(* Logix 5000 project; controller NWGG 1756-L72 rev 35.12; software revision 35.00; part 8 of 19 *)
(* tags used below, declared in another part *)
   _700_AIR_GA : ALIAS FOR I8.3;
   _700_METER : ALIAS FOR I8.2;
   _700_TREAT : ALIAS FOR I7.3;
   _700G_13_CL : ALIAS FOR B21[70].1;
   _700G_13_OP : ALIAS FOR B21[70].0;
   _700G_CLOSE : ALIAS FOR O12.9;
   _700G_OPEN : ALIAS FOR O12.8;
   _701_AIR_GA : ALIAS FOR I8.5;
   _701_FB : ALIAS FOR B21[1].3;
   _701_K_TREA : ALIAS FOR I8.0;
   _701_METER : ALIAS FOR I8.4;
   _701_RB : ALIAS FOR B21[1].4;
   _701_REV_CN : ALIAS FOR C5[3];
   _701_STP : ALIAS FOR B21[1].2;
   _701F_HPB : ALIAS FOR B21[1].0;
   _701F_M : ALIAS FOR O25[10].11;
   _701F_OFF_T : ALIAS FOR T22[1];
   _701G_CLOSE : ALIAS FOR B21[71].13;
   _701G_OPEN : ALIAS FOR B21[71].12;
   _701MR : ALIAS FOR O25[9].7;
   _701R_DELAY : ALIAS FOR T22[2];
   _701R_HPB : ALIAS FOR B21[1].1;
   _701YR : ALIAS FOR I25[1].7;
   _702B : ALIAS FOR B21[2].2;
   _702H_START : ALIAS FOR B21[2].0;
   _702H_STOP : ALIAS FOR B21[2].1;
   _702M : ALIAS FOR O25[9].4;
   _702Y : ALIAS FOR I25[1].4;
   _703B : ALIAS FOR B21[3].2;
   _703H_START : ALIAS FOR B21[3].0;
   _703H_STOP : ALIAS FOR B21[3].1;
   _703M : ALIAS FOR O25[9].14;
   _703Y : ALIAS FOR I25[1].14;
   _704B : ALIAS FOR B21[4].2;
   _704H_START : ALIAS FOR B21[4].0;
   _704H_STOP : ALIAS FOR B21[4].1;
   _704Y : ALIAS FOR I25[0].13;
   _705B : ALIAS FOR B21[5].2;
   _705H_START : ALIAS FOR B21[5].0;
   _705H_STOP : ALIAS FOR B21[5].1;
   _705M : ALIAS FOR O25[10].12;
   _705Y : ALIAS FOR I25[2].12;
   _706B : ALIAS FOR B21[6].2;
   _706H_START : ALIAS FOR B21[6].0;
   _706H_STOP : ALIAS FOR B21[6].1;
   _706M : ALIAS FOR O25[9].11;
   _706Y : ALIAS FOR I25[1].11;
   _707B : ALIAS FOR B21[7].2;
   _707M : ALIAS FOR O25[11].0;
   _707Y : ALIAS FOR I25[3].0;
   _708G_BIN_1 : ALIAS FOR O9.15;
   _709G_BIN_1 : ALIAS FOR O10.15;
   A_HOLD_MB : ALIAS FOR B3[1].3;
   A_HOLD_REL : ALIAS FOR B3[1].5;
   A_STPB_AUT : ALIAS FOR B3[1].1;
   A_TREATER : ALIAS FOR I24[6].8;
   Analog : AI[160];
   CG_19_METR : ALIAS FOR I8.14;
   CONC13_PUM : ALIAS FOR N7[83];
   CONC13_SET1 : ALIAS FOR B21[8].14;
   CONC19_PUM : ALIAS FOR N7[89];
   CONC19_SET : ALIAS FOR B21[9].14;
   CONC_13_NO : ALIAS FOR B21[8].15;
   CONC_19_NO : ALIAS FOR B21[9].15;
   I18_002 : ALIAS FOR I18[2];
   I18_003 : ALIAS FOR I18[3];
   I1_000_Bit00 : ALIAS FOR I1.0;
   I1_000_Bit03 : ALIAS FOR I1.3;
   I1_000_Bit06 : ALIAS FOR I1.6;
   I1_000_Bit09 : ALIAS FOR I1.9;
   I1_000_Bit12 : ALIAS FOR I1.12;
   I24_021_Bit03 : ALIAS FOR I24[21].3;
   I24_021_Bit04 : ALIAS FOR I24[21].4;
   I24_021_Bit05 : ALIAS FOR I24[21].5;
   I24_021_Bit06 : ALIAS FOR I24[21].6;
   I24_021_Bit07 : ALIAS FOR I24[21].7;
   I24_021_Bit08 : ALIAS FOR I24[21].8;
   I2_000_Bit00 : ALIAS FOR I2.0;
   I2_000_Bit03 : ALIAS FOR I2.3;
   I2_000_Bit06 : ALIAS FOR I2.6;
   I2_000_Bit09 : ALIAS FOR I2.9;
   I2_000_Bit12 : ALIAS FOR I2.12;
   I3_000_Bit00 : ALIAS FOR I3.0;
   I3_000_Bit03 : ALIAS FOR I3.3;
   I3_000_Bit06 : ALIAS FOR I3.6;
   I8_000_Bit06 : ALIAS FOR I8.6;
   I8_000_Bit07 : ALIAS FOR I8.7;
   I8_000_Bit08 : ALIAS FOR I8.8;
   I8_000_Bit09 : ALIAS FOR I8.9;
   I8_000_Bit10 : ALIAS FOR I8.10;
   I8_000_Bit11 : ALIAS FOR I8.11;
   MAIN_TIMER : ALIAS FOR T11[0];
   N14 : DINT[84];
   O12_000_Bit10 : ALIAS FOR O12.10;
   O12_000_Bit11 : ALIAS FOR O12.11;
   O12_000_Bit12 : ALIAS FOR O12.12;
   O12_000_Bit13 : ALIAS FOR O12.13;
   O25_008_Bit13 : ALIAS FOR O25[8].13;
   P10_ALARM : ALIAS FOR T4[97];
   P10_ALARM1 : ALIAS FOR T4[99];
   P10_NO_FLO : ALIAS FOR B12[10].3;
   P10_SEC_SE : ALIAS FOR B17[1].10;
   P1_NO_FLOW : ALIAS FOR B12[1].3;
   P2_NO_FLOW : ALIAS FOR B12[2].3;
   P3_NO_FLOW : ALIAS FOR B12[3].3;
   P4_ALARM_N : ALIAS FOR T4[87];
   P4_ALARM_N1 : ALIAS FOR T4[88];
   P4_NO_FLOW : ALIAS FOR B12[4].3;
   P4_SEC_SEL : ALIAS FOR B17[1].4;
   P5_ALARM_N : ALIAS FOR T4[89];
   P5_ALARM_N1 : ALIAS FOR T4[90];
   P5_NO_FLOW : ALIAS FOR B12[5].3;
   P5_SEC_SEL : ALIAS FOR B17[1].5;
   P6_ALARM_N : ALIAS FOR T4[91];
   P6_ALARM_N1 : ALIAS FOR T4[92];
   P6_NO_FLOW : ALIAS FOR B12[6].3;
   P6_SEC_SEL : ALIAS FOR B17[1].6;
   P7_ALARM_N : ALIAS FOR T4[93];
   P7_ALARM_N1 : ALIAS FOR T4[94];
   P7_NO_FLOW : ALIAS FOR B12[7].3;
   P7_SEC_SEL : ALIAS FOR B17[1].7;
   P8_ALARM_N : ALIAS FOR T4[95];
   P8_ALARM_N1 : ALIAS FOR T4[96];
   P8_NO_FLOW : ALIAS FOR B12[8].3;
   P8_SEC_SEL : ALIAS FOR B17[1].8;
   PUMP_NO_FL : ALIAS FOR B12[11].0;
   T11_NO_PAS : ALIAS FOR B17[11].2;
   T12_NO_PAS : ALIAS FOR B17[12].2;
   T13_NO_PAS : ALIAS FOR B17[13].2;
   T13C_CLOSE : ALIAS FOR T22[6];
   T13C_GATE : ALIAS FOR B21[0].0;
   T13C_GATE1 : ALIAS FOR B21[0].1;
   T13C_GATE2 : ALIAS FOR B21[0].3;
   T13C_GATE3 : ALIAS FOR B21[0].4;
   T13C_GATE4 : ALIAS FOR B21[0].5;
   T13C_GATE5 : ALIAS FOR B21[0].6;
   T13C_GATE6 : ALIAS FOR B21[0].7;
   T13C_GATE7 : ALIAS FOR B21[0].8;
   T13C_GATE8 : ALIAS FOR B21[0].9;
   T13C_GATEC : ALIAS FOR B21[0].2;
   T13C_GATET : ALIAS FOR C5[2];
   T13C_TREAT : ALIAS FOR B21[70].10;
   T13C_TRT_M : ALIAS FOR T22[7];
   T13C_TRT_O : ALIAS FOR T22[5];
   T14_NO_PAS : ALIAS FOR B17[14].2;
   T15_NO_PAS : ALIAS FOR B17[15].2;
   T16_NO_PAS : ALIAS FOR B17[16].2;
   T17_NO_PAS : ALIAS FOR B17[17].2;
   T19C_AIR_S : ALIAS FOR B21[71].11;
   T19C_CLOSE1 : ALIAS FOR T22[3];
   T19C_GATE : ALIAS FOR B21[71].0;
   T19C_GATE2 : ALIAS FOR B21[71].3;
   T19C_GATE3 : ALIAS FOR B21[71].4;
   T19C_GATE4 : ALIAS FOR B21[71].5;
   T19C_GATE5 : ALIAS FOR B21[71].6;
   T19C_GATE6 : ALIAS FOR B21[71].7;
   T19C_GATE7 : ALIAS FOR B21[71].8;
   T19C_GATE8 : ALIAS FOR B21[71].9;
   T19C_GATEC : ALIAS FOR B21[71].2;
   T19C_GATET : ALIAS FOR C5[4];
   T19C_TREAT : ALIAS FOR B21[71].10;
   T19C_TRT_M : ALIAS FOR T22[4];
   T19C_TRT_O : ALIAS FOR T22[0];
   T21_NO_PAS : ALIAS FOR B17[21].2;
   T22 : TIMER[100];
   T22_NO_PAS : ALIAS FOR B17[22].2;
   T23_NO_PAS : ALIAS FOR B17[23].2;
   T24_NO_PAS : ALIAS FOR B17[24].2;
   T25_NO_PAS : ALIAS FOR B17[25].2;
   T26_NO_PAS : ALIAS FOR B17[26].2;
   TK11_PUMP : ALIAS FOR N7[70];
   TK12_PUMP : ALIAS FOR N7[71];
   TK13_PUMP : ALIAS FOR N7[72];
   TK14_PUMP : ALIAS FOR N7[73];
   TK15_PUMP : ALIAS FOR N7[74];
   TK16_PUMP : ALIAS FOR N7[75];
   TK17_PUMP : ALIAS FOR N7[76];
   TK21_PUMP : ALIAS FOR N7[77];
   TK22_PUMP : ALIAS FOR N7[78];
   TK23_PUMP : ALIAS FOR N7[79];
   TK24_PUMP : ALIAS FOR N7[80];
   TK25_PUMP : ALIAS FOR N7[81];
   TK26_PUMP : ALIAS FOR N7[82];
(* _2_MAIN, continued *)

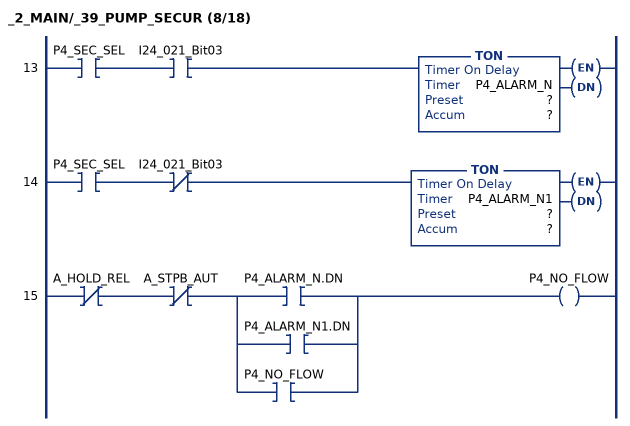
   [picture p142: _2_MAIN/_39_PUMP_SECUR rungs 13-15]
   13: XIC(P4_SEC_SEL)XIC(I24_021_Bit03)TON(P4_ALARM_N,?,?);
   14: XIC(P4_SEC_SEL)XIO(I24_021_Bit03)TON(P4_ALARM_N1,?,?);
   15: XIO(A_HOLD_REL)XIO(A_STPB_AUT)[XIC(P4_ALARM_N.DN) ,XIC(P4_ALARM_N1.DN) ,XIC(P4_NO_FLOW) ]OTE(P4_NO_FLOW);
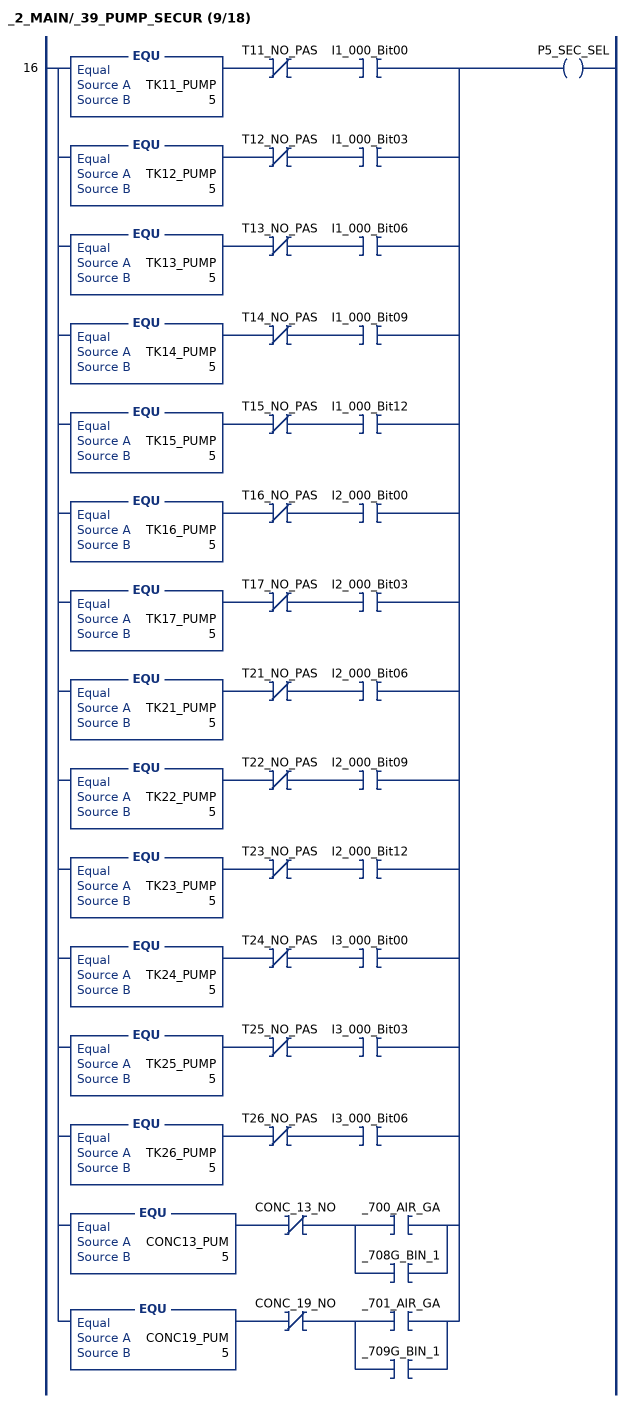
   16: [EQU(TK11_PUMP,5) XIO(T11_NO_PAS) XIC(I1_000_Bit00) ,EQU(TK12_PUMP,5) XIO(T12_NO_PAS) XIC(I1_000_Bit03) ,EQU(TK13_PUMP,5) XIO(T13_NO_PAS) XIC(I1_000_Bit06) ,EQU(TK14_PUMP,5) XIO(T14_NO_PAS) XIC(I1_000_Bit09) ,EQU(TK15_PUMP,5) XIO(T15_NO_PAS) XIC(I1_000_Bit12) ,EQU(TK16_PUMP,5) XIO(T16_NO_PAS) XIC(I2_000_Bit00) ,EQU(TK17_PUMP,5) XIO(T17_NO_PAS) XIC(I2_000_Bit03) ,EQU(TK21_PUMP,5) XIO(T21_NO_PAS) XIC(I2_000_Bit06) ,EQU(TK22_PUMP,5) XIO(T22_NO_PAS) XIC(I2_000_Bit09) ,EQU(TK23_PUMP,5) XIO(T23_NO_PAS) XIC(I2_000_Bit12) ,EQU(TK24_PUMP,5) XIO(T24_NO_PAS) XIC(I3_000_Bit00) ,EQU(TK25_PUMP,5) XIO(T25_NO_PAS) XIC(I3_000_Bit03) ,EQU(TK26_PUMP,5) XIO(T26_NO_PAS) XIC(I3_000_Bit06) ,EQU(CONC13_PUM,5) XIO(CONC_13_NO) [XIC(_700_AIR_GA) ,XIC(_708G_BIN_1) ] ,EQU(CONC19_PUM,5) XIO(CONC_19_NO) [XIC(_701_AIR_GA) ,XIC(_709G_BIN_1) ] ]OTE(P5_SEC_SEL);
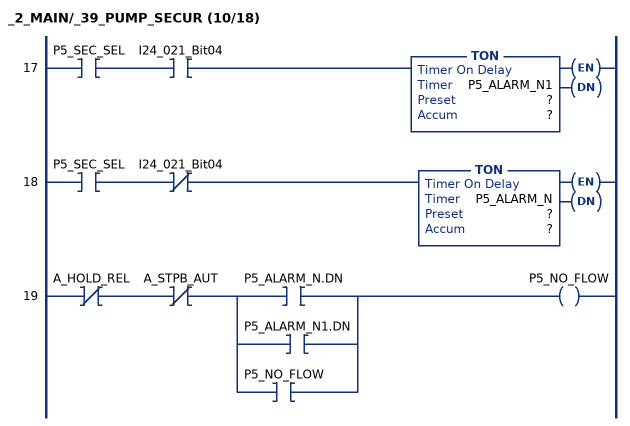
   17: XIC(P5_SEC_SEL)XIC(I24_021_Bit04)TON(P5_ALARM_N1,?,?);
   18: XIC(P5_SEC_SEL)XIO(I24_021_Bit04)TON(P5_ALARM_N,?,?);
   19: XIO(A_HOLD_REL)XIO(A_STPB_AUT)[XIC(P5_ALARM_N.DN) ,XIC(P5_ALARM_N1.DN) ,XIC(P5_NO_FLOW) ]OTE(P5_NO_FLOW);
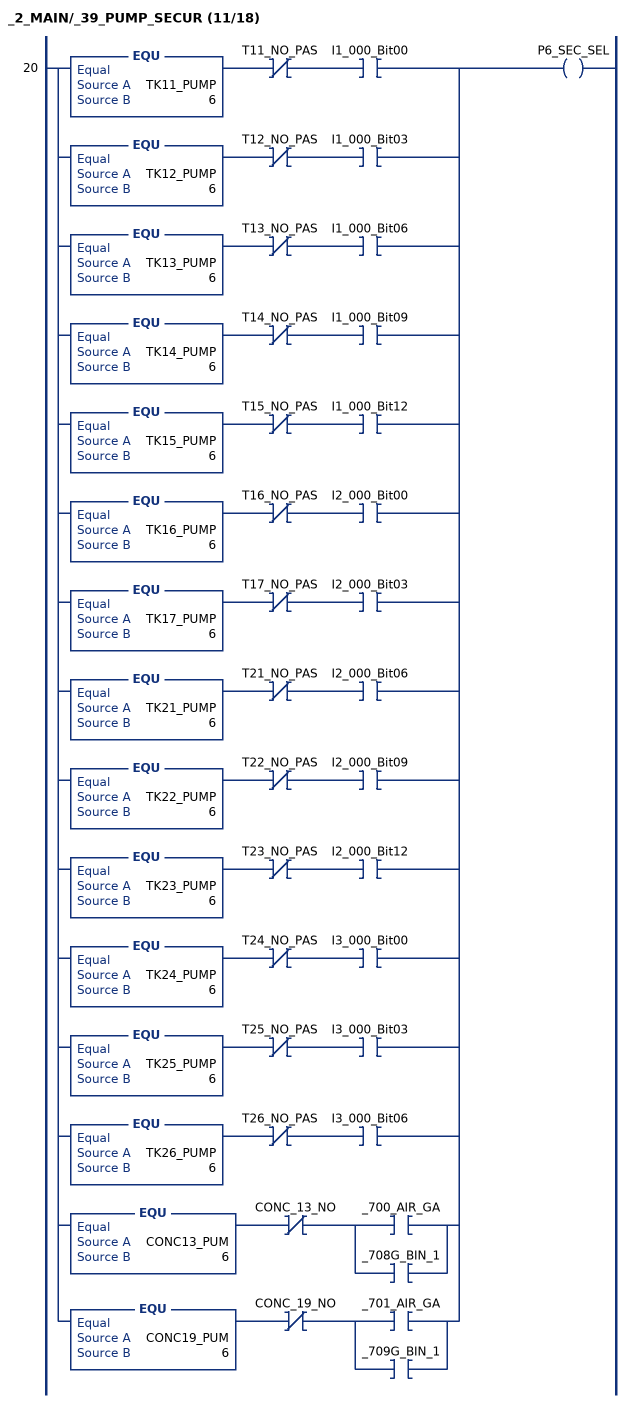
   20: [EQU(TK11_PUMP,6) XIO(T11_NO_PAS) XIC(I1_000_Bit00) ,EQU(TK12_PUMP,6) XIO(T12_NO_PAS) XIC(I1_000_Bit03) ,EQU(TK13_PUMP,6) XIO(T13_NO_PAS) XIC(I1_000_Bit06) ,EQU(TK14_PUMP,6) XIO(T14_NO_PAS) XIC(I1_000_Bit09) ,EQU(TK15_PUMP,6) XIO(T15_NO_PAS) XIC(I1_000_Bit12) ,EQU(TK16_PUMP,6) XIO(T16_NO_PAS) XIC(I2_000_Bit00) ,EQU(TK17_PUMP,6) XIO(T17_NO_PAS) XIC(I2_000_Bit03) ,EQU(TK21_PUMP,6) XIO(T21_NO_PAS) XIC(I2_000_Bit06) ,EQU(TK22_PUMP,6) XIO(T22_NO_PAS) XIC(I2_000_Bit09) ,EQU(TK23_PUMP,6) XIO(T23_NO_PAS) XIC(I2_000_Bit12) ,EQU(TK24_PUMP,6) XIO(T24_NO_PAS) XIC(I3_000_Bit00) ,EQU(TK25_PUMP,6) XIO(T25_NO_PAS) XIC(I3_000_Bit03) ,EQU(TK26_PUMP,6) XIO(T26_NO_PAS) XIC(I3_000_Bit06) ,EQU(CONC13_PUM,6) XIO(CONC_13_NO) [XIC(_700_AIR_GA) ,XIC(_708G_BIN_1) ] ,EQU(CONC19_PUM,6) XIO(CONC_19_NO) [XIC(_701_AIR_GA) ,XIC(_709G_BIN_1) ] ]OTE(P6_SEC_SEL);
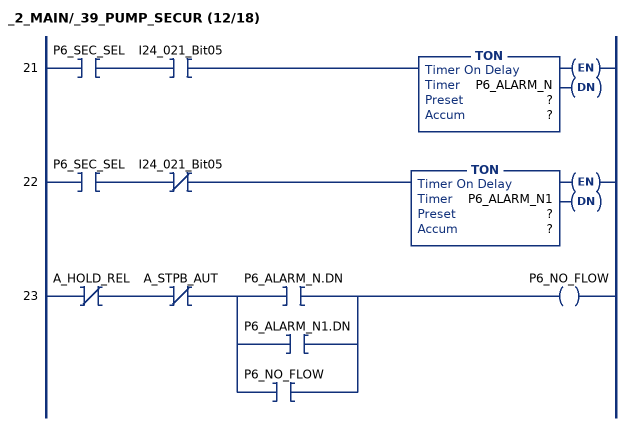
   21: XIC(P6_SEC_SEL)XIC(I24_021_Bit05)TON(P6_ALARM_N,?,?);
   22: XIC(P6_SEC_SEL)XIO(I24_021_Bit05)TON(P6_ALARM_N1,?,?);
   23: XIO(A_HOLD_REL)XIO(A_STPB_AUT)[XIC(P6_ALARM_N.DN) ,XIC(P6_ALARM_N1.DN) ,XIC(P6_NO_FLOW) ]OTE(P6_NO_FLOW);
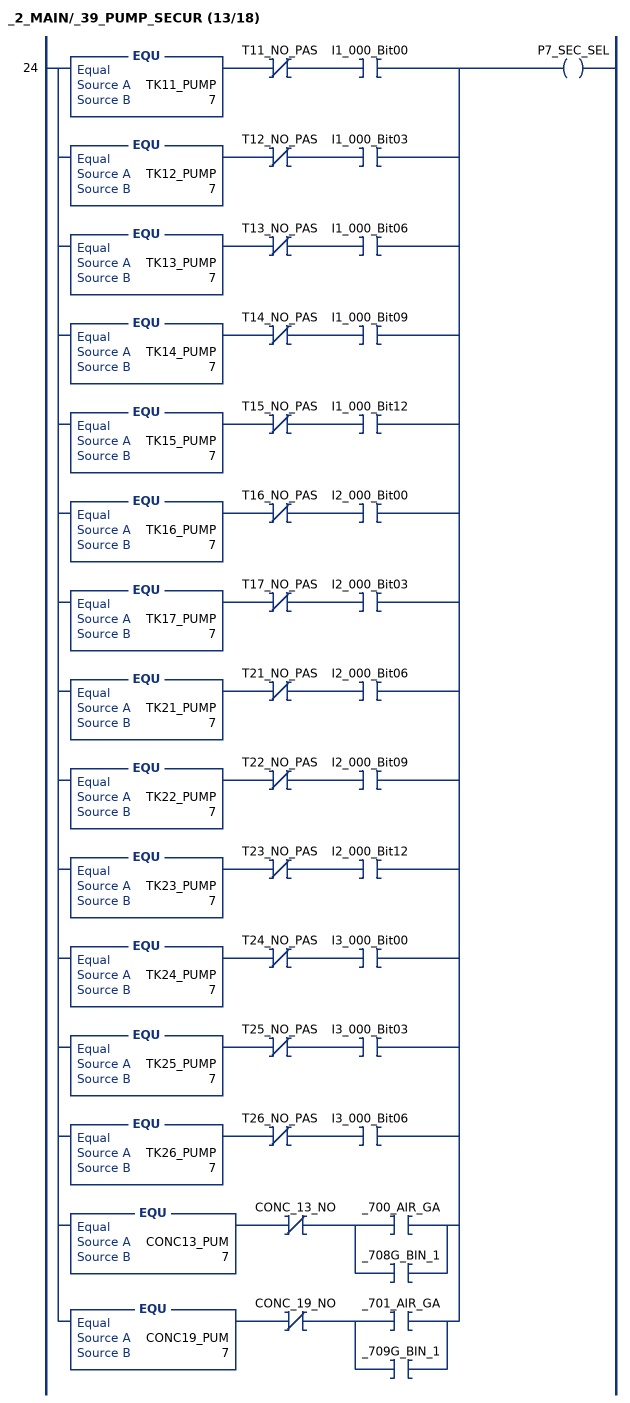
   24: [EQU(TK11_PUMP,7) XIO(T11_NO_PAS) XIC(I1_000_Bit00) ,EQU(TK12_PUMP,7) XIO(T12_NO_PAS) XIC(I1_000_Bit03) ,EQU(TK13_PUMP,7) XIO(T13_NO_PAS) XIC(I1_000_Bit06) ,EQU(TK14_PUMP,7) XIO(T14_NO_PAS) XIC(I1_000_Bit09) ,EQU(TK15_PUMP,7) XIO(T15_NO_PAS) XIC(I1_000_Bit12) ,EQU(TK16_PUMP,7) XIO(T16_NO_PAS) XIC(I2_000_Bit00) ,EQU(TK17_PUMP,7) XIO(T17_NO_PAS) XIC(I2_000_Bit03) ,EQU(TK21_PUMP,7) XIO(T21_NO_PAS) XIC(I2_000_Bit06) ,EQU(TK22_PUMP,7) XIO(T22_NO_PAS) XIC(I2_000_Bit09) ,EQU(TK23_PUMP,7) XIO(T23_NO_PAS) XIC(I2_000_Bit12) ,EQU(TK24_PUMP,7) XIO(T24_NO_PAS) XIC(I3_000_Bit00) ,EQU(TK25_PUMP,7) XIO(T25_NO_PAS) XIC(I3_000_Bit03) ,EQU(TK26_PUMP,7) XIO(T26_NO_PAS) XIC(I3_000_Bit06) ,EQU(CONC13_PUM,7) XIO(CONC_13_NO) [XIC(_700_AIR_GA) ,XIC(_708G_BIN_1) ] ,EQU(CONC19_PUM,7) XIO(CONC_19_NO) [XIC(_701_AIR_GA) ,XIC(_709G_BIN_1) ] ]OTE(P7_SEC_SEL);
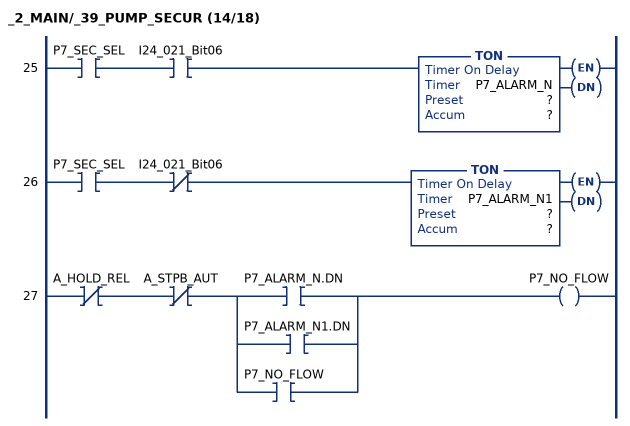
   25: XIC(P7_SEC_SEL)XIC(I24_021_Bit06)TON(P7_ALARM_N,?,?);
   26: XIC(P7_SEC_SEL)XIO(I24_021_Bit06)TON(P7_ALARM_N1,?,?);
   27: XIO(A_HOLD_REL)XIO(A_STPB_AUT)[XIC(P7_ALARM_N.DN) ,XIC(P7_ALARM_N1.DN) ,XIC(P7_NO_FLOW) ]OTE(P7_NO_FLOW);
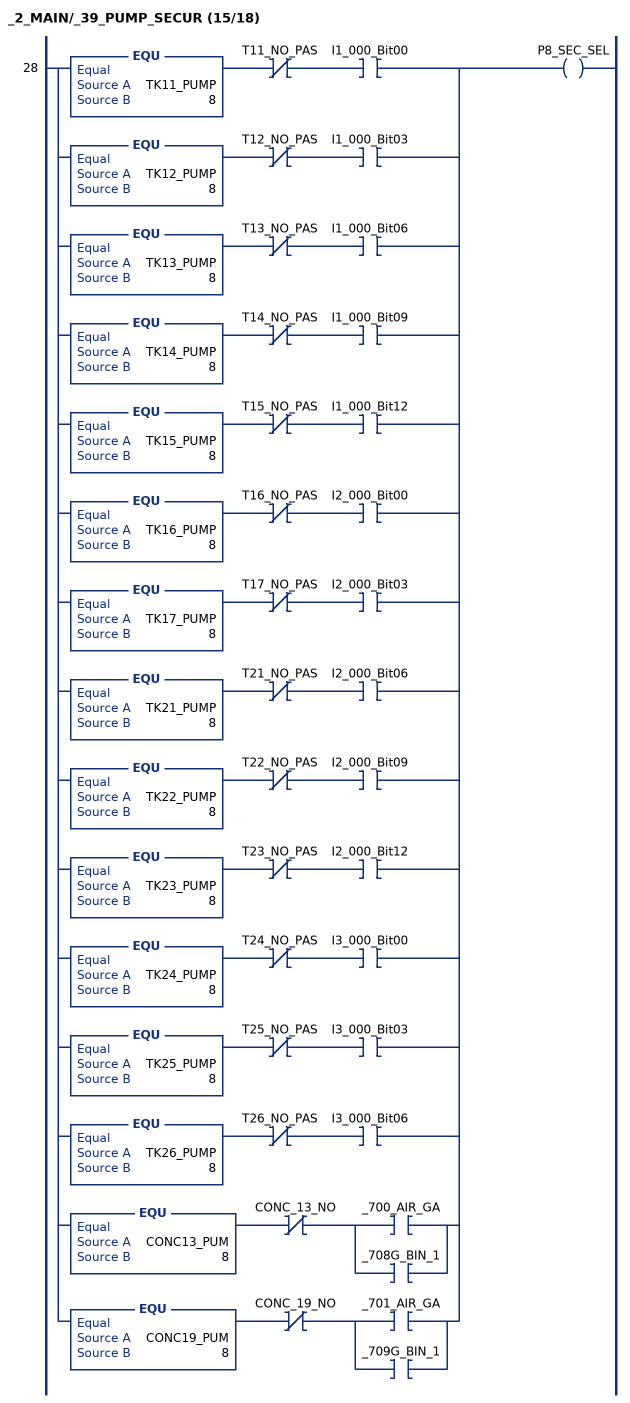
   28: [EQU(TK11_PUMP,8) XIO(T11_NO_PAS) XIC(I1_000_Bit00) ,EQU(TK12_PUMP,8) XIO(T12_NO_PAS) XIC(I1_000_Bit03) ,EQU(TK13_PUMP,8) XIO(T13_NO_PAS) XIC(I1_000_Bit06) ,EQU(TK14_PUMP,8) XIO(T14_NO_PAS) XIC(I1_000_Bit09) ,EQU(TK15_PUMP,8) XIO(T15_NO_PAS) XIC(I1_000_Bit12) ,EQU(TK16_PUMP,8) XIO(T16_NO_PAS) XIC(I2_000_Bit00) ,EQU(TK17_PUMP,8) XIO(T17_NO_PAS) XIC(I2_000_Bit03) ,EQU(TK21_PUMP,8) XIO(T21_NO_PAS) XIC(I2_000_Bit06) ,EQU(TK22_PUMP,8) XIO(T22_NO_PAS) XIC(I2_000_Bit09) ,EQU(TK23_PUMP,8) XIO(T23_NO_PAS) XIC(I2_000_Bit12) ,EQU(TK24_PUMP,8) XIO(T24_NO_PAS) XIC(I3_000_Bit00) ,EQU(TK25_PUMP,8) XIO(T25_NO_PAS) XIC(I3_000_Bit03) ,EQU(TK26_PUMP,8) XIO(T26_NO_PAS) XIC(I3_000_Bit06) ,EQU(CONC13_PUM,8) XIO(CONC_13_NO) [XIC(_700_AIR_GA) ,XIC(_708G_BIN_1) ] ,EQU(CONC19_PUM,8) XIO(CONC_19_NO) [XIC(_701_AIR_GA) ,XIC(_709G_BIN_1) ] ]OTE(P8_SEC_SEL);
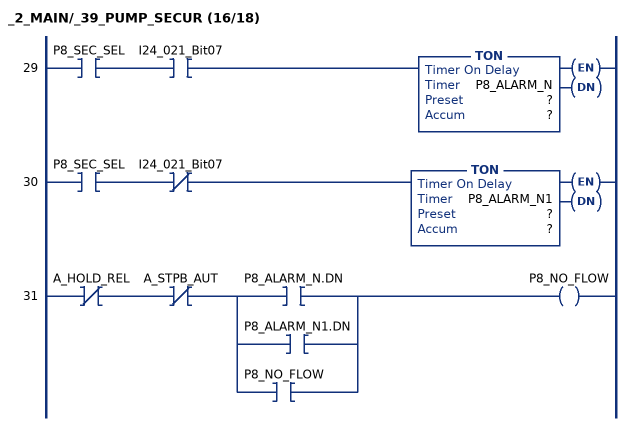
   29: XIC(P8_SEC_SEL)XIC(I24_021_Bit07)TON(P8_ALARM_N,?,?);
   30: XIC(P8_SEC_SEL)XIO(I24_021_Bit07)TON(P8_ALARM_N1,?,?);
   31: XIO(A_HOLD_REL)XIO(A_STPB_AUT)[XIC(P8_ALARM_N.DN) ,XIC(P8_ALARM_N1.DN) ,XIC(P8_NO_FLOW) ]OTE(P8_NO_FLOW);
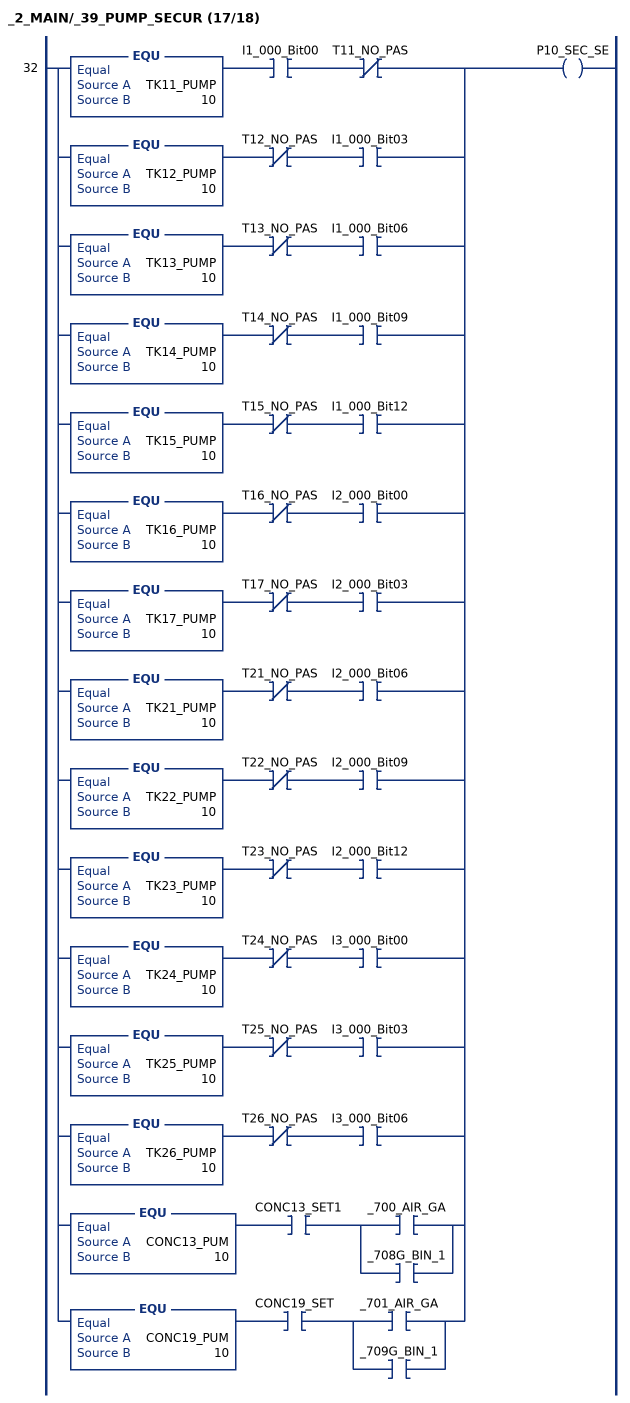
   32: [EQU(TK11_PUMP,10) XIC(I1_000_Bit00) XIO(T11_NO_PAS) ,EQU(TK12_PUMP,10) XIO(T12_NO_PAS) XIC(I1_000_Bit03) ,EQU(TK13_PUMP,10) XIO(T13_NO_PAS) XIC(I1_000_Bit06) ,EQU(TK14_PUMP,10) XIO(T14_NO_PAS) XIC(I1_000_Bit09) ,EQU(TK15_PUMP,10) XIO(T15_NO_PAS) XIC(I1_000_Bit12) ,EQU(TK16_PUMP,10) XIO(T16_NO_PAS) XIC(I2_000_Bit00) ,EQU(TK17_PUMP,10) XIO(T17_NO_PAS) XIC(I2_000_Bit03) ,EQU(TK21_PUMP,10) XIO(T21_NO_PAS) XIC(I2_000_Bit06) ,EQU(TK22_PUMP,10) XIO(T22_NO_PAS) XIC(I2_000_Bit09) ,EQU(TK23_PUMP,10) XIO(T23_NO_PAS) XIC(I2_000_Bit12) ,EQU(TK24_PUMP,10) XIO(T24_NO_PAS) XIC(I3_000_Bit00) ,EQU(TK25_PUMP,10) XIO(T25_NO_PAS) XIC(I3_000_Bit03) ,EQU(TK26_PUMP,10) XIO(T26_NO_PAS) XIC(I3_000_Bit06) ,EQU(CONC13_PUM,10) XIC(CONC13_SET1) [XIC(_700_AIR_GA) ,XIC(_708G_BIN_1) ] ,EQU(CONC19_PUM,10) XIC(CONC19_SET) [XIC(_701_AIR_GA) ,XIC(_709G_BIN_1) ] ]OTE(P10_SEC_SE);
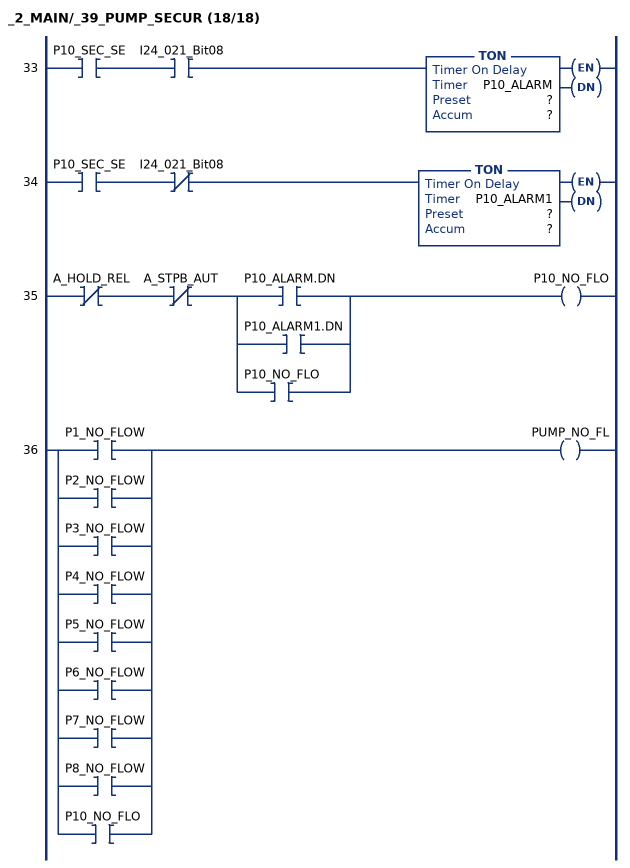
   33: XIC(P10_SEC_SE)XIC(I24_021_Bit08)TON(P10_ALARM,?,?);
   34: XIC(P10_SEC_SE)XIO(I24_021_Bit08)TON(P10_ALARM1,?,?);
   35: XIO(A_HOLD_REL)XIO(A_STPB_AUT)[XIC(P10_ALARM.DN) ,XIC(P10_ALARM1.DN) ,XIC(P10_NO_FLO) ]OTE(P10_NO_FLO);
   36: [XIC(P1_NO_FLOW) ,XIC(P2_NO_FLOW) ,XIC(P3_NO_FLOW) ,XIC(P4_NO_FLOW) ,XIC(P5_NO_FLOW) ,XIC(P6_NO_FLOW) ,XIC(P7_NO_FLOW) ,XIC(P8_NO_FLOW) ,XIC(P10_NO_FLO) ]OTE(PUMP_NO_FL);
END_ROUTINE

ROUTINE _40_TANK_13_19   (* ladder *)
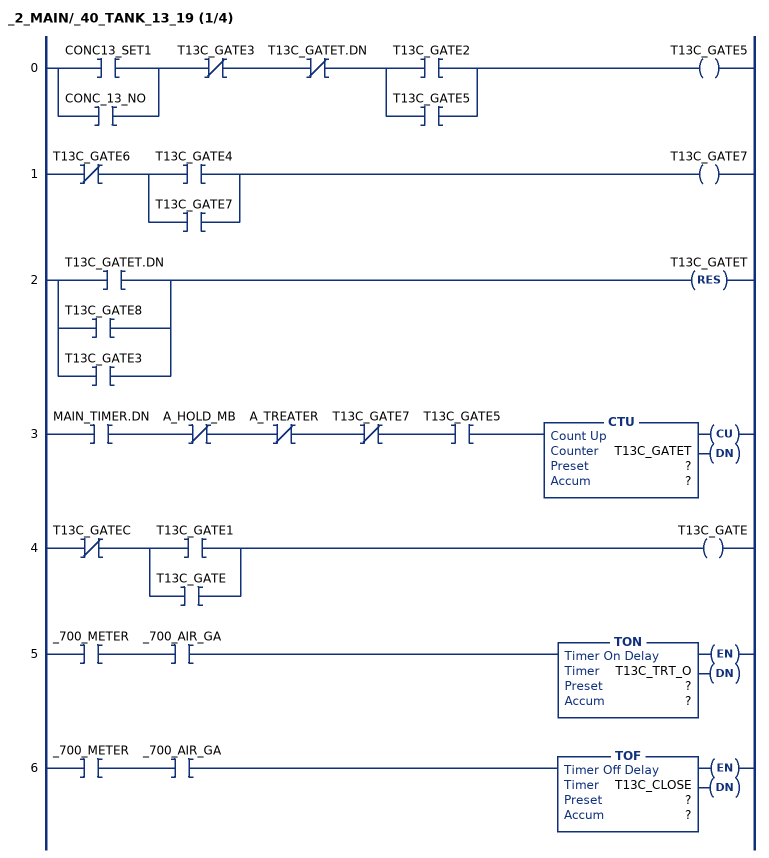
   0: [XIC(CONC13_SET1) ,XIC(CONC_13_NO) ]XIO(T13C_GATE3)XIO(T13C_GATET.DN)[XIC(T13C_GATE2) ,XIC(T13C_GATE5) ]OTE(T13C_GATE5);
   1: XIO(T13C_GATE6)[XIC(T13C_GATE4) ,XIC(T13C_GATE7) ]OTE(T13C_GATE7);
   2: [XIC(T13C_GATET.DN) ,XIC(T13C_GATE8) ,XIC(T13C_GATE3) ]RES(T13C_GATET);
   3: XIC(MAIN_TIMER.DN)XIO(A_HOLD_MB)XIO(A_TREATER)XIO(T13C_GATE7)XIC(T13C_GATE5)CTU(T13C_GATET,?,?);
   4: XIO(T13C_GATEC)[XIC(T13C_GATE1) ,XIC(T13C_GATE) ]OTE(T13C_GATE);
   5: XIC(_700_METER)XIC(_700_AIR_GA)TON(T13C_TRT_O,?,?);
   6: XIC(_700_METER)XIC(_700_AIR_GA)TOF(T13C_CLOSE,?,?);
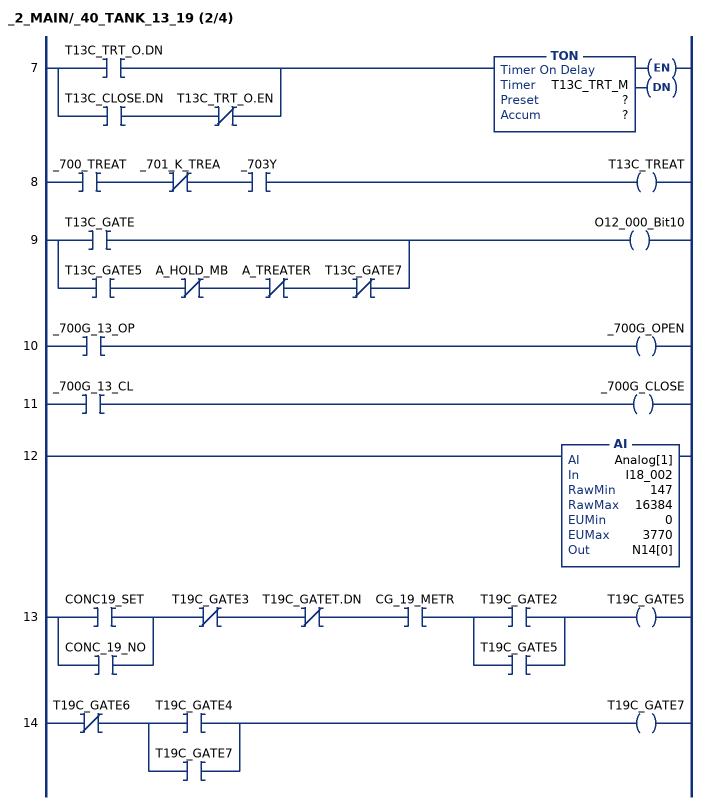
   7: [XIC(T13C_TRT_O.DN) ,XIC(T13C_CLOSE.DN) XIO(T13C_TRT_O.EN) ]TON(T13C_TRT_M,?,?);
   8: XIC(_700_TREAT)XIO(_701_K_TREA)XIC(_703Y)OTE(T13C_TREAT);
   9: [XIC(T13C_GATE) ,XIC(T13C_GATE5) XIO(A_HOLD_MB) XIO(A_TREATER) XIO(T13C_GATE7) ]OTE(O12_000_Bit10);
   10: XIC(_700G_13_OP)OTE(_700G_OPEN);
   11: XIC(_700G_13_CL)OTE(_700G_CLOSE);
   12: AI(Analog[1],I18_002,147,16384,0,3770,N14[0]);
   13: [XIC(CONC19_SET) ,XIC(CONC_19_NO) ]XIO(T19C_GATE3)XIO(T19C_GATET.DN)XIC(CG_19_METR)[XIC(T19C_GATE2) ,XIC(T19C_GATE5) ]OTE(T19C_GATE5);
   14: XIO(T19C_GATE6)[XIC(T19C_GATE4) ,XIC(T19C_GATE7) ]OTE(T19C_GATE7);
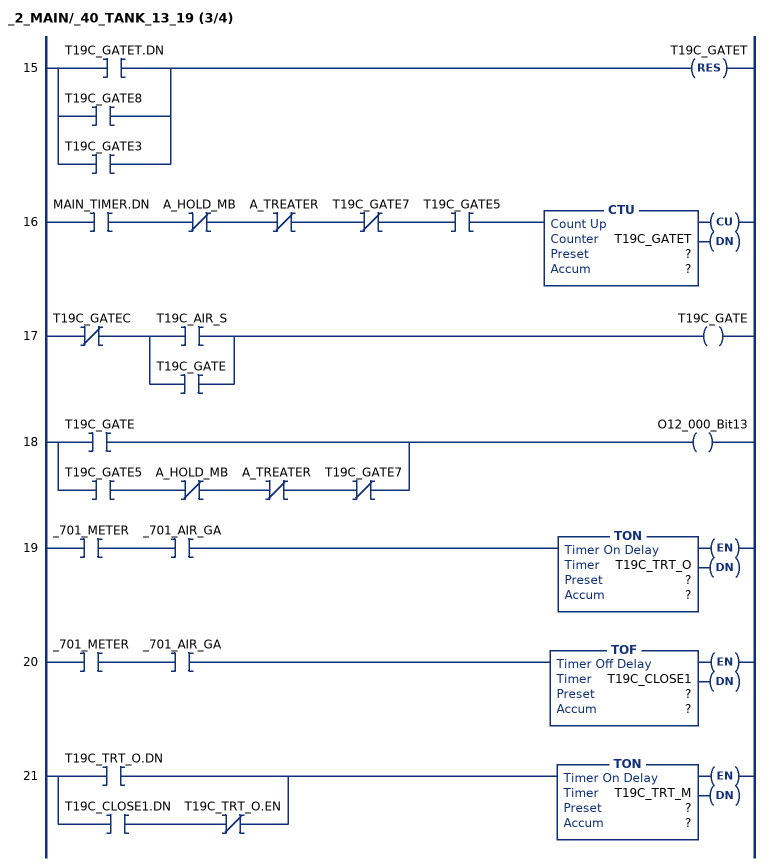
   15: [XIC(T19C_GATET.DN) ,XIC(T19C_GATE8) ,XIC(T19C_GATE3) ]RES(T19C_GATET);
   16: XIC(MAIN_TIMER.DN)XIO(A_HOLD_MB)XIO(A_TREATER)XIO(T19C_GATE7)XIC(T19C_GATE5)CTU(T19C_GATET,?,?);
   17: XIO(T19C_GATEC)[XIC(T19C_AIR_S) ,XIC(T19C_GATE) ]OTE(T19C_GATE);
   18: [XIC(T19C_GATE) ,XIC(T19C_GATE5) XIO(A_HOLD_MB) XIO(A_TREATER) XIO(T19C_GATE7) ]OTE(O12_000_Bit13);
   19: XIC(_701_METER)XIC(_701_AIR_GA)TON(T19C_TRT_O,?,?);
   20: XIC(_701_METER)XIC(_701_AIR_GA)TOF(T19C_CLOSE1,?,?);
   21: [XIC(T19C_TRT_O.DN) ,XIC(T19C_CLOSE1.DN) XIO(T19C_TRT_O.EN) ]TON(T19C_TRT_M,?,?);
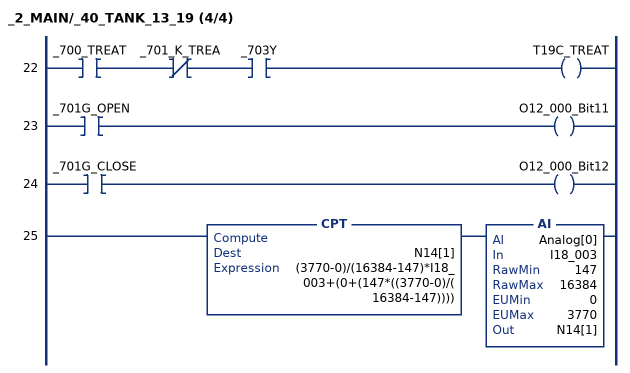
   22: XIC(_700_TREAT)XIO(_701_K_TREA)XIC(_703Y)OTE(T19C_TREAT);
   23: XIC(_701G_OPEN)OTE(O12_000_Bit11);
   24: XIC(_701G_CLOSE)OTE(O12_000_Bit12);
   25: CPT(N14[1],(3770-0)/(16384-147)*I18_003+(0+(147*((3770-0)/(16384-147)))))AI(Analog[0],I18_003,147,16384,0,3770,N14[1]);
END_ROUTINE

ROUTINE _41_CONC_BINS   (* ladder *)
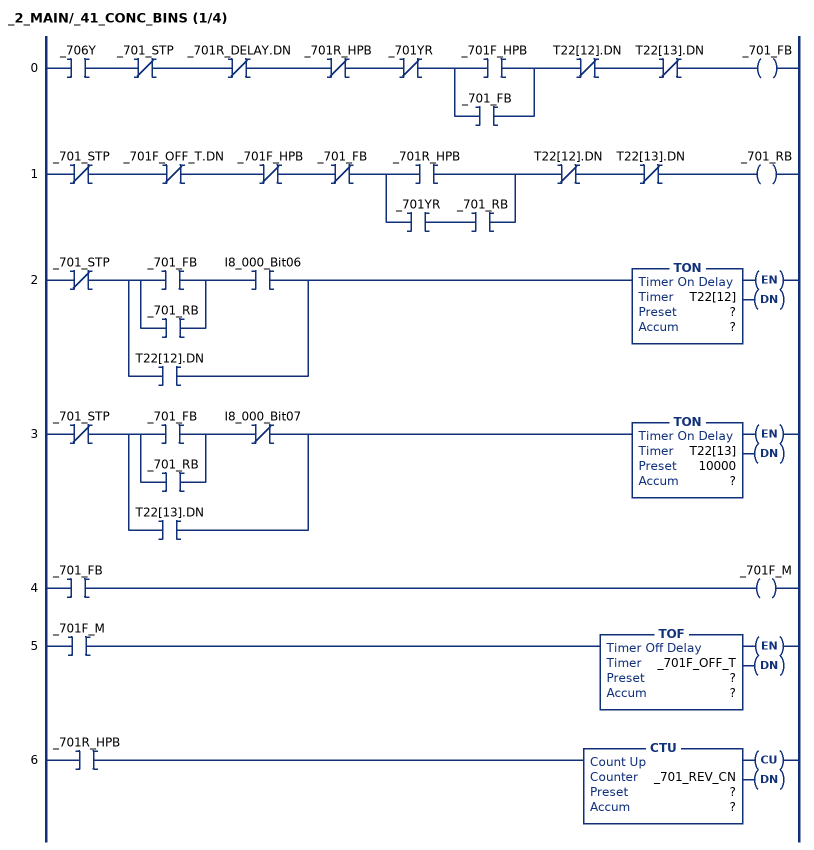
   0: XIC(_706Y)XIO(_701_STP)XIO(_701R_DELAY.DN)XIO(_701R_HPB)XIO(_701YR)[XIC(_701F_HPB) ,XIC(_701_FB) ]XIO(T22[12].DN)XIO(T22[13].DN)OTE(_701_FB);
   1: XIO(_701_STP)XIO(_701F_OFF_T.DN)XIO(_701F_HPB)XIO(_701_FB)[XIC(_701R_HPB) ,XIC(_701YR) XIC(_701_RB) ]XIO(T22[12].DN)XIO(T22[13].DN)OTE(_701_RB);
   2: XIO(_701_STP)[[XIC(_701_FB) ,XIC(_701_RB) ] XIC(I8_000_Bit06) ,XIC(T22[12].DN) ]TON(T22[12],?,?);
   3: XIO(_701_STP)[[XIC(_701_FB) ,XIC(_701_RB) ] XIO(I8_000_Bit07) ,XIC(T22[13].DN) ]TON(T22[13],?,?);
   4: XIC(_701_FB)OTE(_701F_M);
   5: XIC(_701F_M)TOF(_701F_OFF_T,?,?);
   6: XIC(_701R_HPB)CTU(_701_REV_CN,?,?);
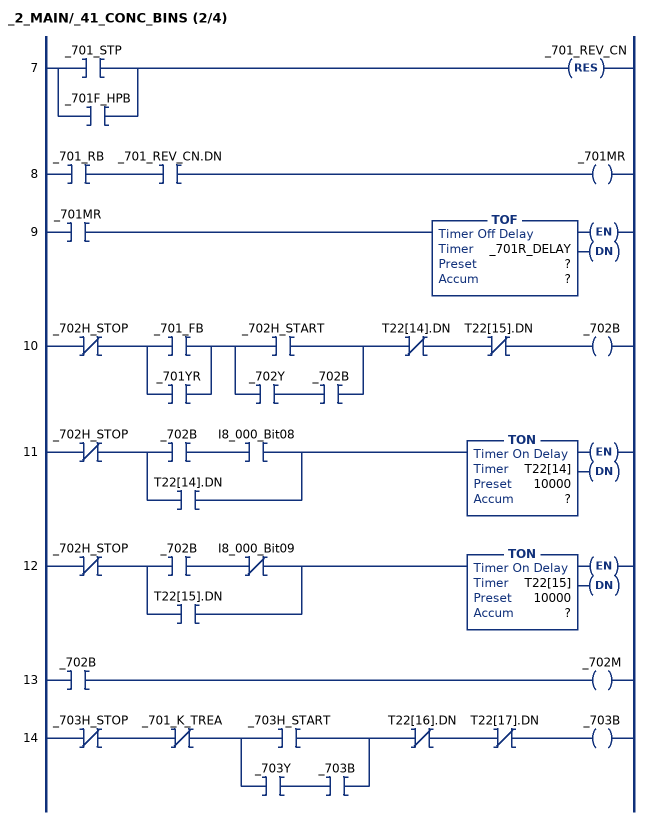
   7: [XIC(_701_STP) ,XIC(_701F_HPB) ]RES(_701_REV_CN);
   8: XIC(_701_RB)XIC(_701_REV_CN.DN)OTE(_701MR);
   9: XIC(_701MR)TOF(_701R_DELAY,?,?);
   10: XIO(_702H_STOP)[XIC(_701_FB) ,XIC(_701YR) ][XIC(_702H_START) ,XIC(_702Y) XIC(_702B) ]XIO(T22[14].DN)XIO(T22[15].DN)OTE(_702B);
   11: XIO(_702H_STOP)[XIC(_702B) XIC(I8_000_Bit08) ,XIC(T22[14].DN) ]TON(T22[14],?,?);
   12: XIO(_702H_STOP)[XIC(_702B) XIO(I8_000_Bit09) ,XIC(T22[15].DN) ]TON(T22[15],?,?);
   13: XIC(_702B)OTE(_702M);
   14: XIO(_703H_STOP)XIO(_701_K_TREA)[XIC(_703H_START) ,XIC(_703Y) XIC(_703B) ]XIO(T22[16].DN)XIO(T22[17].DN)OTE(_703B);
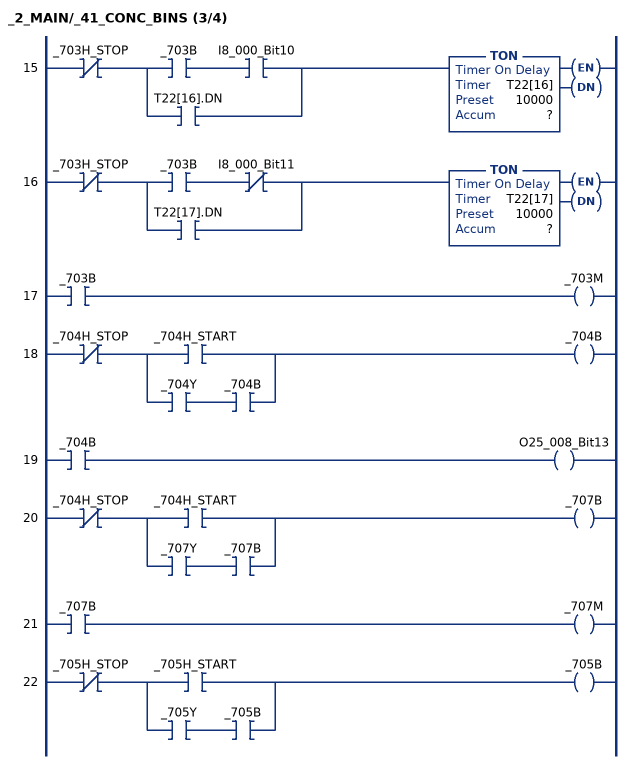
   15: XIO(_703H_STOP)[XIC(_703B) XIC(I8_000_Bit10) ,XIC(T22[16].DN) ]TON(T22[16],?,?);
   16: XIO(_703H_STOP)[XIC(_703B) XIO(I8_000_Bit11) ,XIC(T22[17].DN) ]TON(T22[17],?,?);
   17: XIC(_703B)OTE(_703M);
   18: XIO(_704H_STOP)[XIC(_704H_START) ,XIC(_704Y) XIC(_704B) ]OTE(_704B);
   19: XIC(_704B)OTE(O25_008_Bit13);
   20: XIO(_704H_STOP)[XIC(_704H_START) ,XIC(_707Y) XIC(_707B) ]OTE(_707B);
   21: XIC(_707B)OTE(_707M);
   22: XIO(_705H_STOP)[XIC(_705H_START) ,XIC(_705Y) XIC(_705B) ]OTE(_705B);
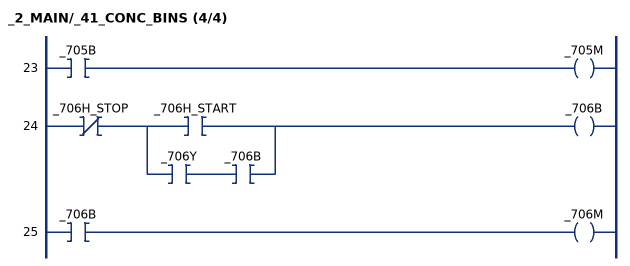
   23: XIC(_705B)OTE(_705M);
   24: XIO(_706H_STOP)[XIC(_706H_START) ,XIC(_706Y) XIC(_706B) ]OTE(_706B);
   25: XIC(_706B)OTE(_706M);
END_ROUTINE
